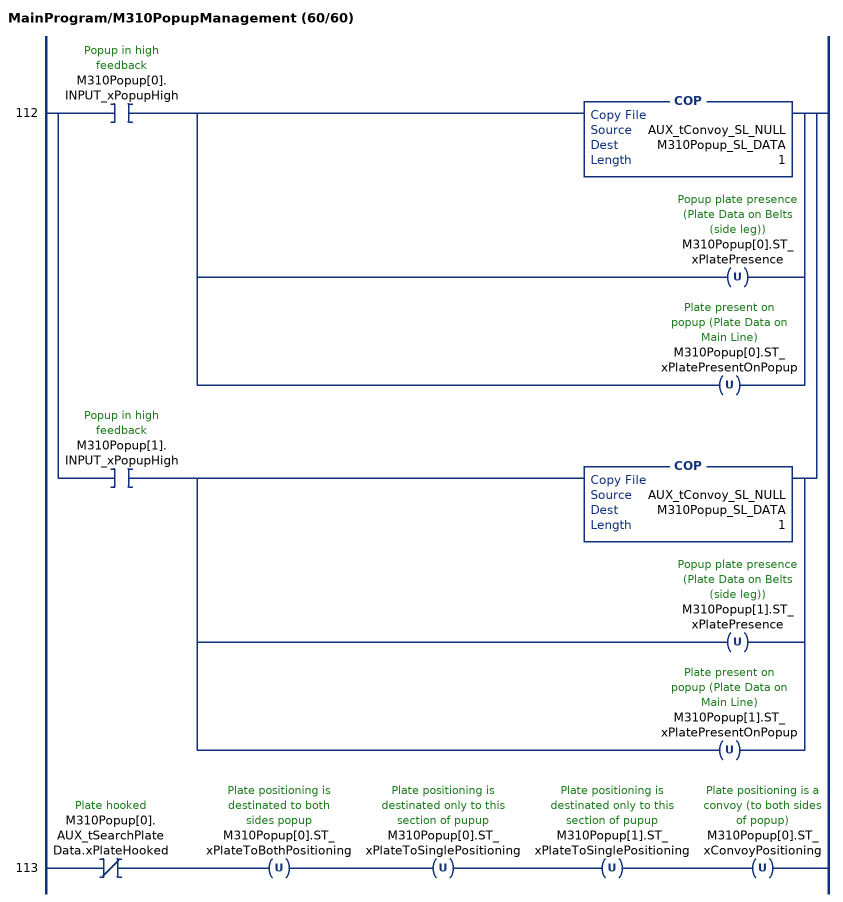
   112: [XIC(M310Popup[0].INPUT_xPopupHigh) [COP(AUX_tConvoy_SL_NULL,M310Popup_SL_DATA,1) ,OTU(M310Popup[0].ST_xPlatePresence) ,OTU(M310Popup[0].ST_xPlatePresentOnPopup) ] ,XIC(M310Popup[1].INPUT_xPopupHigh) [COP(AUX_tConvoy_SL_NULL,M310Popup_SL_DATA,1) ,OTU(M310Popup[1].ST_xPlatePresence) ,OTU(M310Popup[1].ST_xPlatePresentOnPopup) ] ];
   113: XIO(M310Popup[0].AUX_tSearchPlateData.xPlateHooked)OTU(M310Popup[0].ST_xPlateToBothPositioning)OTU(M310Popup[0].ST_xPlateToSinglePositioning)OTU(M310Popup[1].ST_xPlateToSinglePositioning)OTU(M310Popup[0].ST_xConvoyPositioning);
END_ROUTINE

ROUTINE M311_Alarm   (* ladder *)
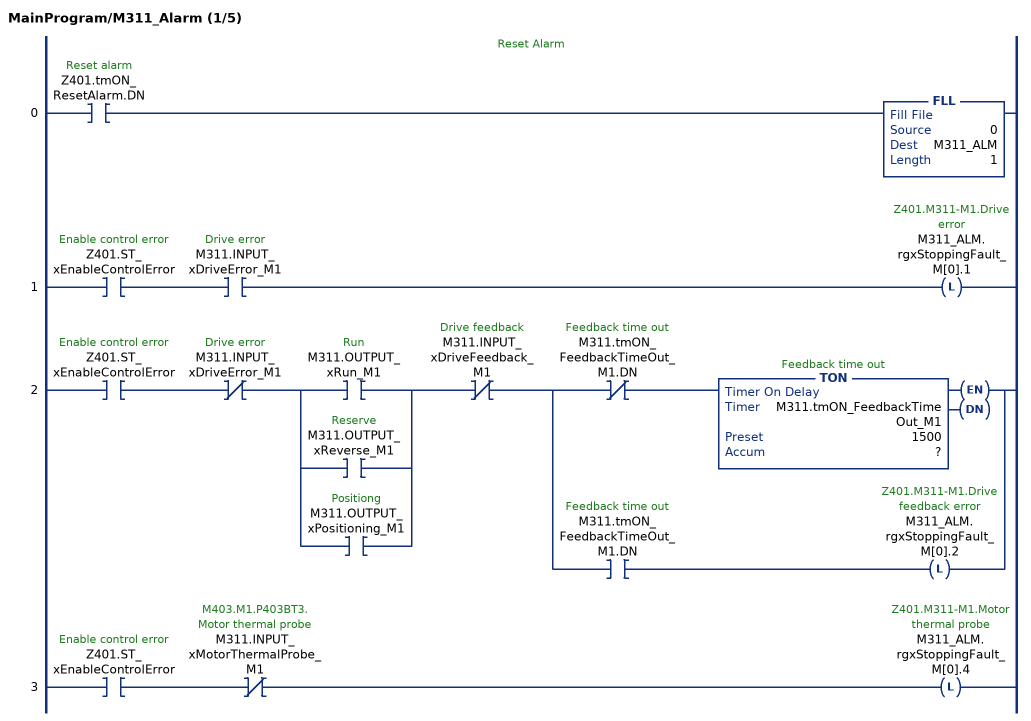
   // Reset Alarm
   0: XIC(Z401.tmON_ResetAlarm.DN)FLL(0,M311_ALM,1);
   1: XIC(Z401.ST_xEnableControlError)XIC(M311.INPUT_xDriveError_M1)OTL(M311_ALM.rgxStoppingFault_M[0].1);
   2: XIC(Z401.ST_xEnableControlError)XIO(M311.INPUT_xDriveError_M1)[XIC(M311.OUTPUT_xRun_M1) ,XIC(M311.OUTPUT_xReverse_M1) ,XIC(M311.OUTPUT_xPositioning_M1) ]XIO(M311.INPUT_xDriveFeedback_M1)[XIO(M311.tmON_FeedbackTimeOut_M1.DN) TON(M311.tmON_FeedbackTimeOut_M1,?,?) ,XIC(M311.tmON_FeedbackTimeOut_M1.DN) OTL(M311_ALM.rgxStoppingFault_M[0].2) ];
   3: XIC(Z401.ST_xEnableControlError)XIO(M311.INPUT_xMotorThermalProbe_M1)OTL(M311_ALM.rgxStoppingFault_M[0].4);
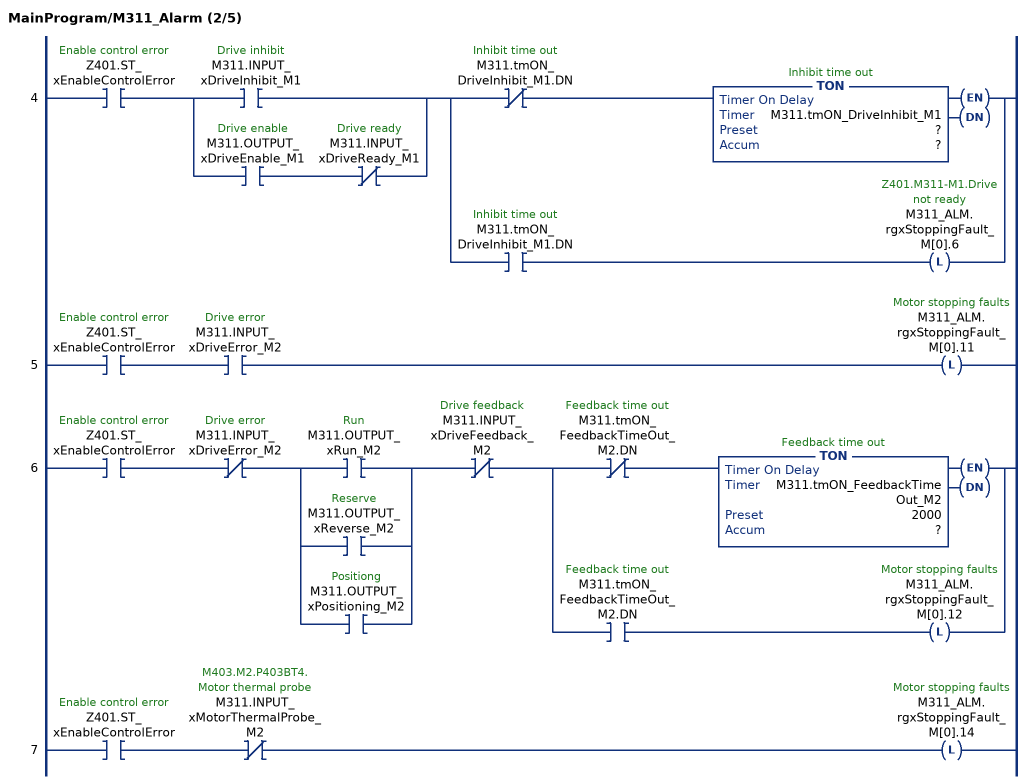
   4: XIC(Z401.ST_xEnableControlError)[XIC(M311.INPUT_xDriveInhibit_M1) ,XIC(M311.OUTPUT_xDriveEnable_M1) XIO(M311.INPUT_xDriveReady_M1) ][XIO(M311.tmON_DriveInhibit_M1.DN) TON(M311.tmON_DriveInhibit_M1,?,?) ,XIC(M311.tmON_DriveInhibit_M1.DN) OTL(M311_ALM.rgxStoppingFault_M[0].6) ];
   5: XIC(Z401.ST_xEnableControlError)XIC(M311.INPUT_xDriveError_M2)OTL(M311_ALM.rgxStoppingFault_M[0].11);
   6: XIC(Z401.ST_xEnableControlError)XIO(M311.INPUT_xDriveError_M2)[XIC(M311.OUTPUT_xRun_M2) ,XIC(M311.OUTPUT_xReverse_M2) ,XIC(M311.OUTPUT_xPositioning_M2) ]XIO(M311.INPUT_xDriveFeedback_M2)[XIO(M311.tmON_FeedbackTimeOut_M2.DN) TON(M311.tmON_FeedbackTimeOut_M2,?,?) ,XIC(M311.tmON_FeedbackTimeOut_M2.DN) OTL(M311_ALM.rgxStoppingFault_M[0].12) ];
   7: XIC(Z401.ST_xEnableControlError)XIO(M311.INPUT_xMotorThermalProbe_M2)OTL(M311_ALM.rgxStoppingFault_M[0].14);
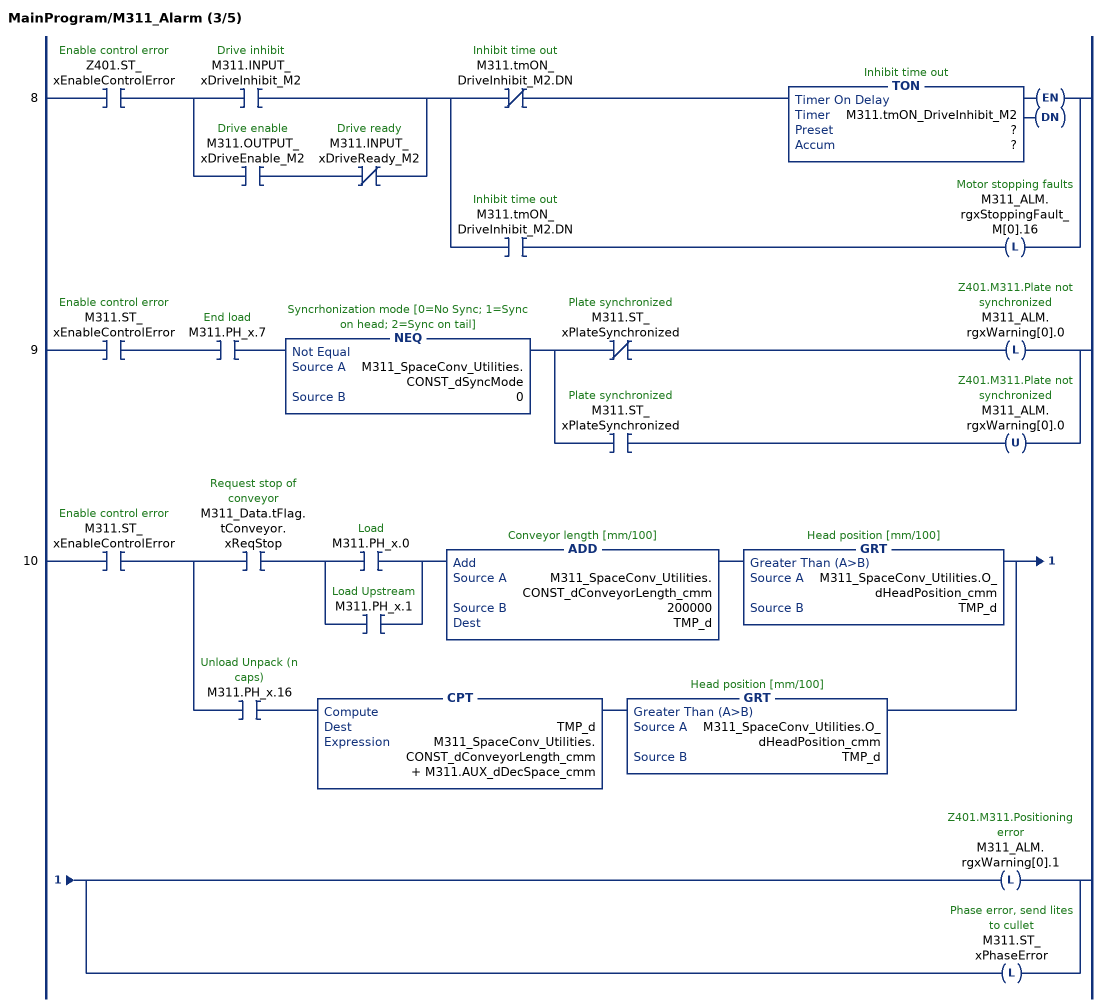
   8: XIC(Z401.ST_xEnableControlError)[XIC(M311.INPUT_xDriveInhibit_M2) ,XIC(M311.OUTPUT_xDriveEnable_M2) XIO(M311.INPUT_xDriveReady_M2) ][XIO(M311.tmON_DriveInhibit_M2.DN) TON(M311.tmON_DriveInhibit_M2,?,?) ,XIC(M311.tmON_DriveInhibit_M2.DN) OTL(M311_ALM.rgxStoppingFault_M[0].16) ];
   9: XIC(M311.ST_xEnableControlError)XIC(M311.PH_x.7)NEQ(M311_SpaceConv_Utilities.CONST_dSyncMode,0)[XIO(M311.ST_xPlateSynchronized) OTL(M311_ALM.rgxWarning[0].0) ,XIC(M311.ST_xPlateSynchronized) OTU(M311_ALM.rgxWarning[0].0) ];
   10: XIC(M311.ST_xEnableControlError)[XIC(M311_Data.tFlag.tConveyor.xReqStop) [XIC(M311.PH_x.0) ,XIC(M311.PH_x.1) ] ADD(M311_SpaceConv_Utilities.CONST_dConveyorLength_cmm,200000,TMP_d) GRT(M311_SpaceConv_Utilities.O_dHeadPosition_cmm,TMP_d) ,XIC(M311.PH_x.16) CPT(TMP_d,M311_SpaceConv_Utilities.CONST_dConveyorLength_cmm + M311.AUX_dDecSpace_cmm) GRT(M311_SpaceConv_Utilities.O_dHeadPosition_cmm,TMP_d) ][OTL(M311_ALM.rgxWarning[0].1) ,OTL(M311.ST_xPhaseError) ];
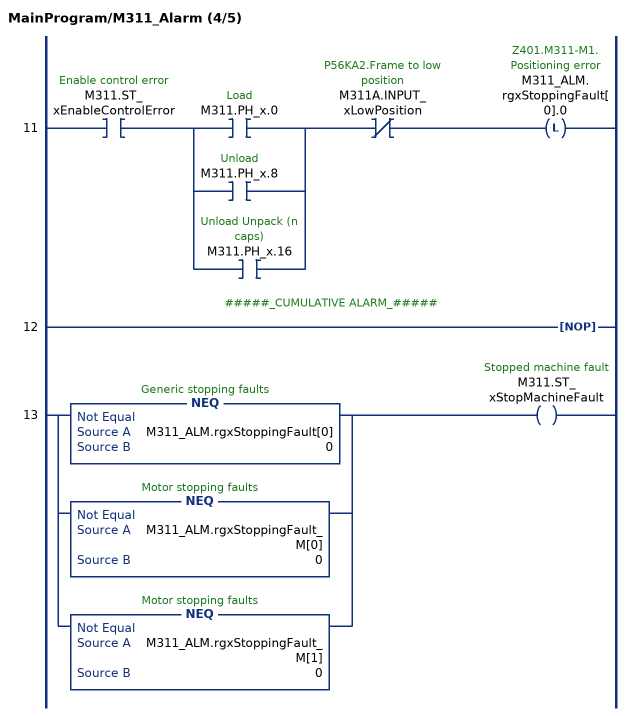
   11: XIC(M311.ST_xEnableControlError)[XIC(M311.PH_x.0) ,XIC(M311.PH_x.8) ,XIC(M311.PH_x.16) ]XIO(M311A.INPUT_xLowPosition)OTL(M311_ALM.rgxStoppingFault[0].0);
   // #####_CUMULATIVE ALARM_#####
   12: NOP();
   13: [NEQ(M311_ALM.rgxStoppingFault[0],0) ,NEQ(M311_ALM.rgxStoppingFault_M[0],0) ,NEQ(M311_ALM.rgxStoppingFault_M[1],0) ]OTE(M311.ST_xStopMachineFault);
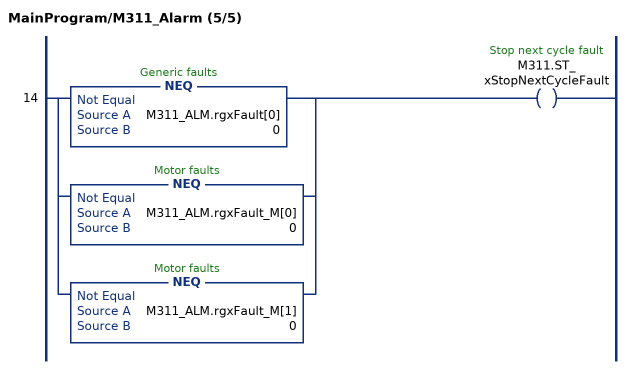
   14: [NEQ(M311_ALM.rgxFault[0],0) ,NEQ(M311_ALM.rgxFault_M[0],0) ,NEQ(M311_ALM.rgxFault_M[1],0) ]OTE(M311.ST_xStopNextCycleFault);
END_ROUTINE

ROUTINE M311_Logic   (* ladder *)
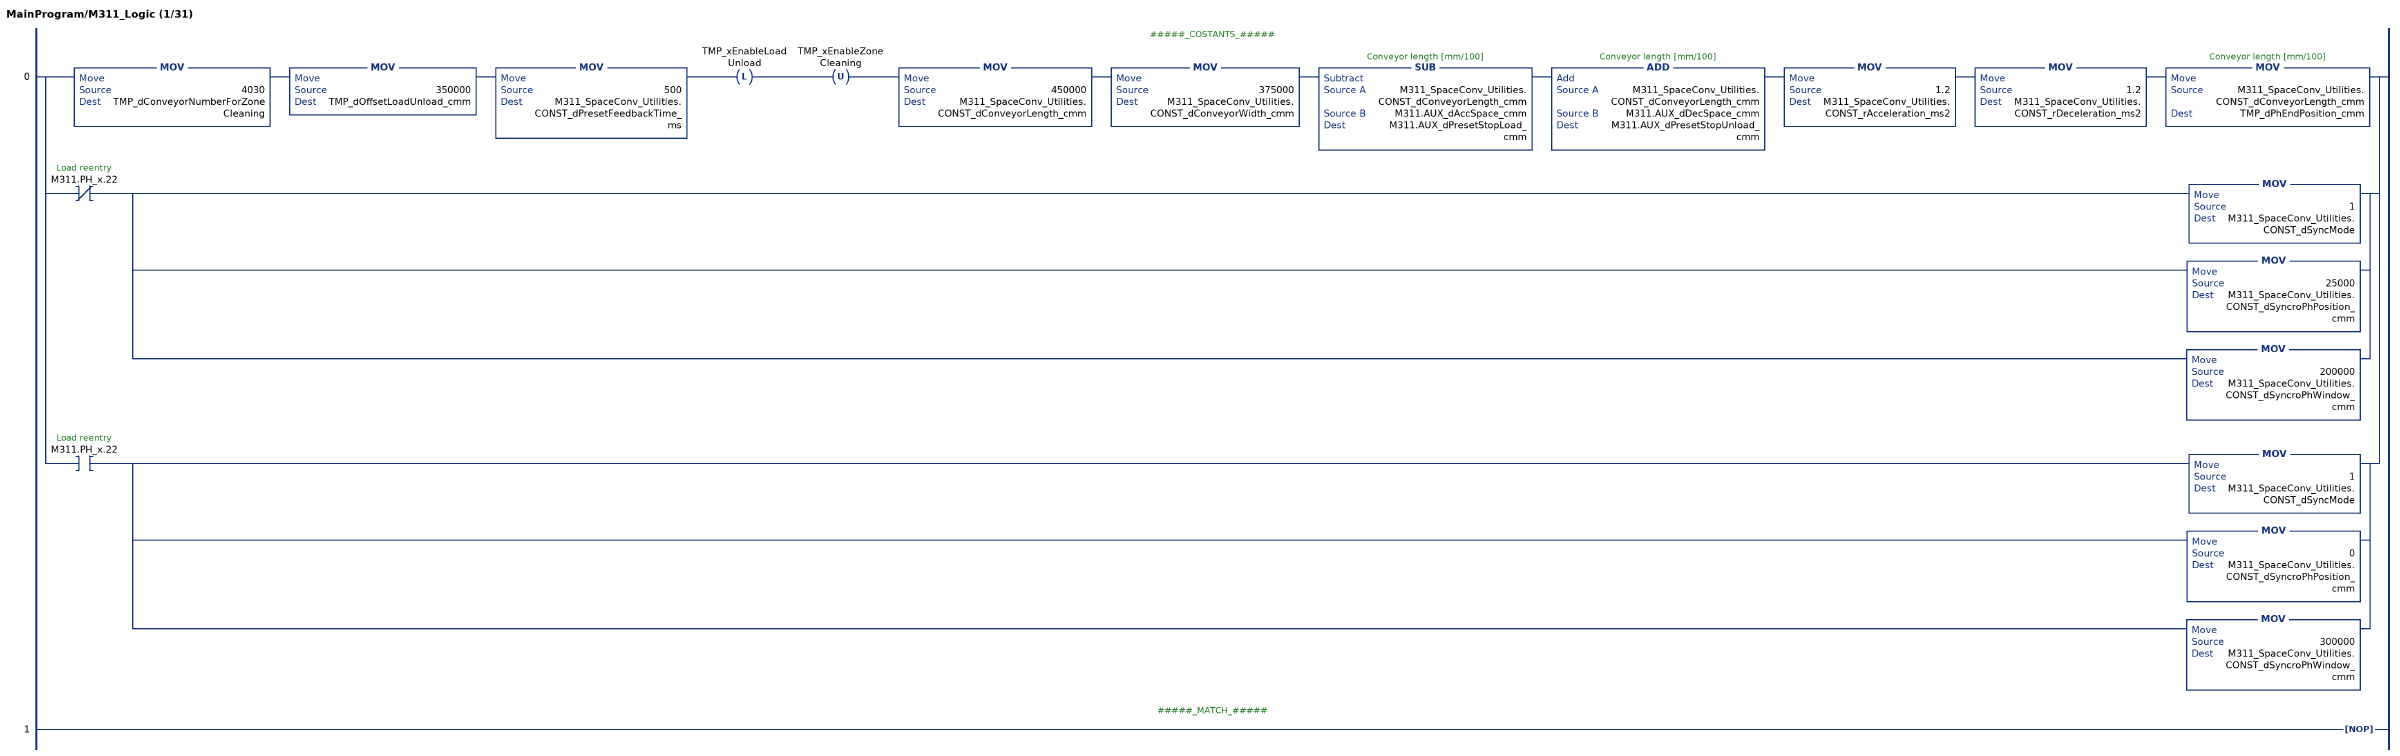
   // #####_COSTANTS_#####
   0: [MOV(4030,TMP_dConveyorNumberForZoneCleaning) MOV(350000,TMP_dOffsetLoadUnload_cmm) MOV(500,M311_SpaceConv_Utilities.CONST_dPresetFeedbackTime_ms) OTL(TMP_xEnableLoadUnload) OTU(TMP_xEnableZoneCleaning) MOV(450000,M311_SpaceConv_Utilities.CONST_dConveyorLength_cmm) MOV(375000,M311_SpaceConv_Utilities.CONST_dConveyorWidth_cmm) SUB(M311_SpaceConv_Utilities.CONST_dConveyorLength_cmm,M311.AUX_dAccSpace_cmm,M311.AUX_dPresetStopLoad_cmm) ADD(M311_SpaceConv_Utilities.CONST_dConveyorLength_cmm,M311.AUX_dDecSpace_cmm,M311.AUX_dPresetStopUnload_cmm) MOV(1.2,M311_SpaceConv_Utilities.CONST_rAcceleration_ms2) MOV(1.2,M311_SpaceConv_Utilities.CONST_rDeceleration_ms2) MOV(M311_SpaceConv_Utilities.CONST_dConveyorLength_cmm,TMP_dPhEndPosition_cmm) ,XIO(M311.PH_x.22) [MOV(1,M311_SpaceConv_Utilities.CONST_dSyncMode) ,MOV(25000,M311_SpaceConv_Utilities.CONST_dSyncroPhPosition_cmm) ,MOV(200000,M311_SpaceConv_Utilities.CONST_dSyncroPhWindow_cmm) ] ,XIC(M311.PH_x.22) [MOV(1,M311_SpaceConv_Utilities.CONST_dSyncMode) ,MOV(0,M311_SpaceConv_Utilities.CONST_dSyncroPhPosition_cmm) ,MOV(300000,M311_SpaceConv_Utilities.CONST_dSyncroPhWindow_cmm) ] ];
   // #####_MATCH_#####
   1: NOP();
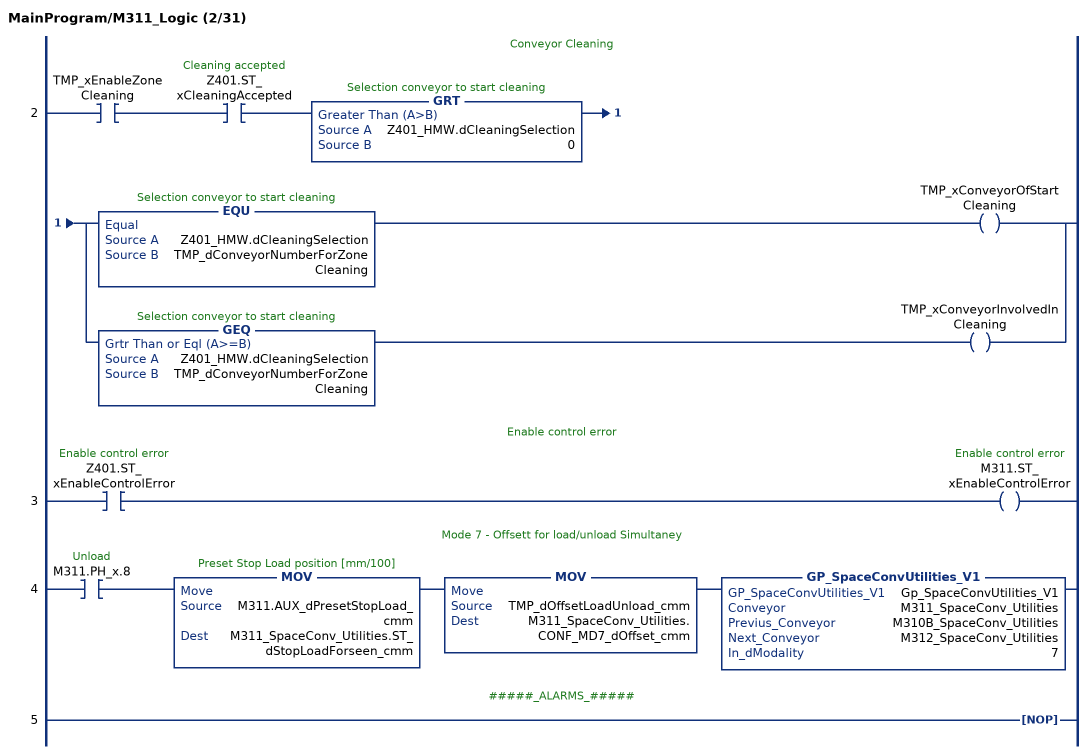
   // Conveyor Cleaning
   2: XIC(TMP_xEnableZoneCleaning)XIC(Z401.ST_xCleaningAccepted)GRT(Z401_HMW.dCleaningSelection,0)[EQU(Z401_HMW.dCleaningSelection,TMP_dConveyorNumberForZoneCleaning) OTE(TMP_xConveyorOfStartCleaning) ,GEQ(Z401_HMW.dCleaningSelection,TMP_dConveyorNumberForZoneCleaning) OTE(TMP_xConveyorInvolvedInCleaning) ];
   // Enable control error
   3: XIC(Z401.ST_xEnableControlError)OTE(M311.ST_xEnableControlError);
   // Mode 7 - Offsett for load/unload Simultaney
   4: XIC(M311.PH_x.8)MOV(M311.AUX_dPresetStopLoad_cmm,M311_SpaceConv_Utilities.ST_dStopLoadForseen_cmm)MOV(TMP_dOffsetLoadUnload_cmm,M311_SpaceConv_Utilities.CONF_MD7_dOffset_cmm)GP_SpaceConvUtilities_V1(Gp_SpaceConvUtilities_V1,M311_SpaceConv_Utilities,M310B_SpaceConv_Utilities,M312_SpaceConv_Utilities,7);
   // #####_ALARMS_#####
   5: NOP();
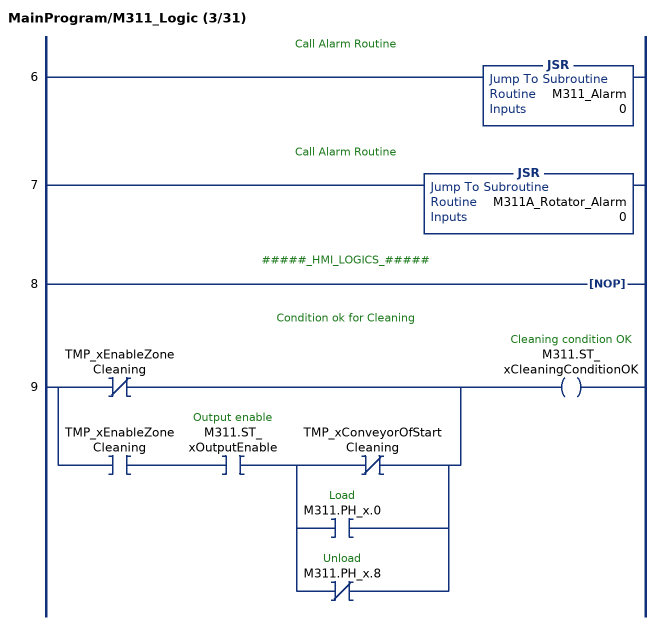
   // Call Alarm Routine
   6: JSR(M311_Alarm,0);
   // Call Alarm Routine
   7: JSR(M311A_Rotator_Alarm,0);
   // #####_HMI_LOGICS_#####
   8: NOP();
   // Condition ok for Cleaning
   9: [XIO(TMP_xEnableZoneCleaning) ,XIC(TMP_xEnableZoneCleaning) XIC(M311.ST_xOutputEnable) [XIO(TMP_xConveyorOfStartCleaning) ,XIC(M311.PH_x.0) ,XIO(M311.PH_x.8) ] ]OTE(M311.ST_xCleaningConditionOK);
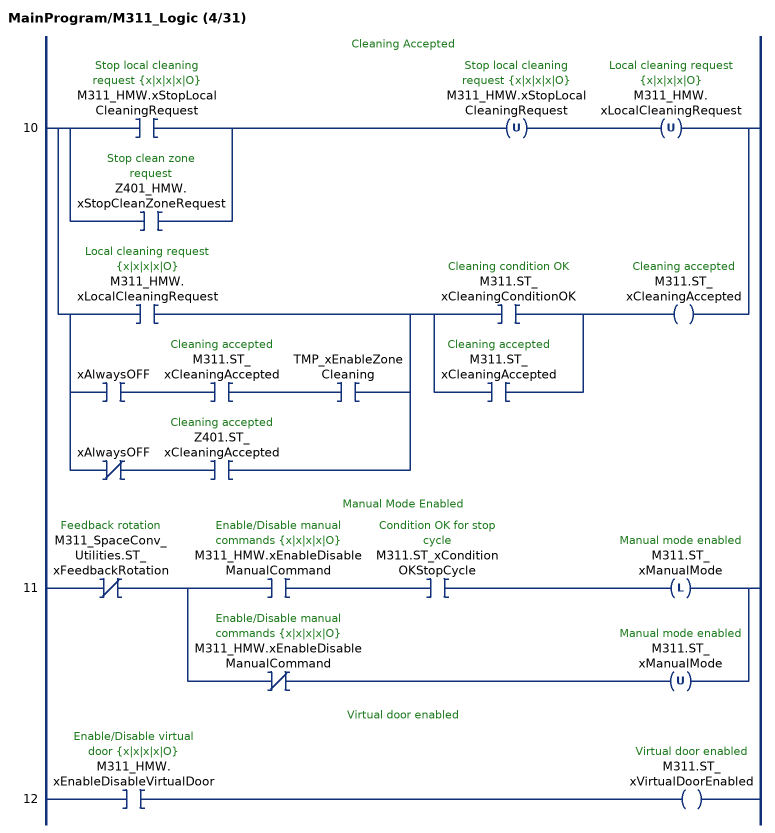
   // Cleaning Accepted
   10: [[XIC(M311_HMW.xStopLocalCleaningRequest) ,XIC(Z401_HMW.xStopCleanZoneRequest) ] OTU(M311_HMW.xStopLocalCleaningRequest) OTU(M311_HMW.xLocalCleaningRequest) ,[XIC(M311_HMW.xLocalCleaningRequest) ,XIC(xAlwaysOFF) XIC(M311.ST_xCleaningAccepted) XIC(TMP_xEnableZoneCleaning) ,XIO(xAlwaysOFF) XIC(Z401.ST_xCleaningAccepted) ] [XIC(M311.ST_xCleaningConditionOK) ,XIC(M311.ST_xCleaningAccepted) ] OTE(M311.ST_xCleaningAccepted) ];
   // Manual Mode Enabled
   11: XIO(M311_SpaceConv_Utilities.ST_xFeedbackRotation)[XIC(M311_HMW.xEnableDisableManualCommand) XIC(M311.ST_xConditionOKStopCycle) OTL(M311.ST_xManualMode) ,XIO(M311_HMW.xEnableDisableManualCommand) OTU(M311.ST_xManualMode) ];
   // Virtual door enabled
   12: XIC(M311_HMW.xEnableDisableVirtualDoor)OTE(M311.ST_xVirtualDoorEnabled);
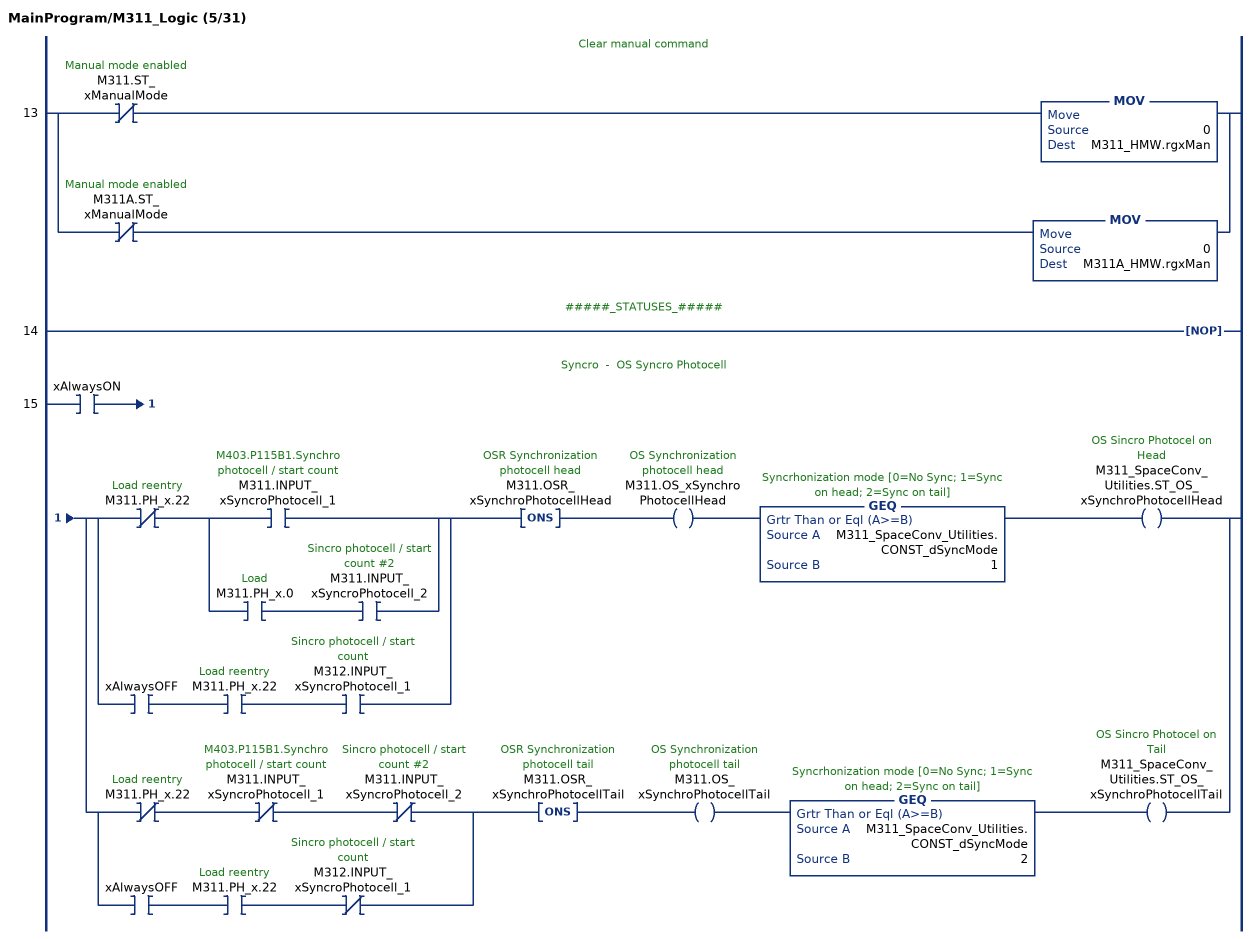
   // Clear manual command
   13: [XIO(M311.ST_xManualMode) MOV(0,M311_HMW.rgxMan) ,XIO(M311A.ST_xManualMode) MOV(0,M311A_HMW.rgxMan) ];
   // #####_STATUSES_#####
   14: NOP();
   // Syncro  -  OS Syncro Photocell
   15: XIC(xAlwaysON)[[XIO(M311.PH_x.22) [XIC(M311.INPUT_xSyncroPhotocell_1) ,XIC(M311.PH_x.0) XIC(M311.INPUT_xSyncroPhotocell_2) ] ,XIC(xAlwaysOFF) XIC(M311.PH_x.22) XIC(M312.INPUT_xSyncroPhotocell_1) ] ONS(M311.OSR_xSynchroPhotocellHead) OTE(M311.OS_xSynchroPhotocellHead) GEQ(M311_SpaceConv_Utilities.CONST_dSyncMode,1) OTE(M311_SpaceConv_Utilities.ST_OS_xSynchroPhotocellHead) ,[XIO(M311.PH_x.22) XIO(M311.INPUT_xSyncroPhotocell_1) XIO(M311.INPUT_xSyncroPhotocell_2) ,XIC(xAlwaysOFF) XIC(M311.PH_x.22) XIO(M312.INPUT_xSyncroPhotocell_1) ] ONS(M311.OSR_xSynchroPhotocellTail) OTE(M311.OS_xSynchroPhotocellTail) GEQ(M311_SpaceConv_Utilities.CONST_dSyncMode,2) OTE(M311_SpaceConv_Utilities.ST_OS_xSynchroPhotocellTail) ];
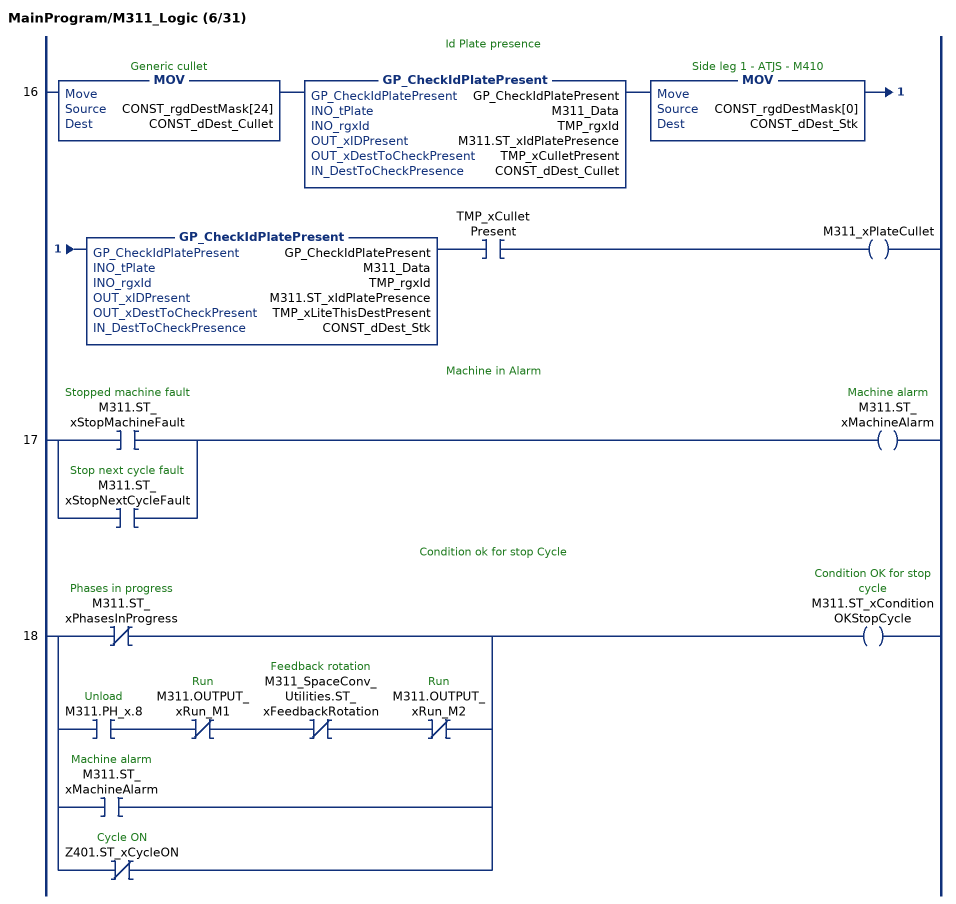
   // Id Plate presence
   16: MOV(CONST_rgdDestMask[24],CONST_dDest_Cullet)GP_CheckIdPlatePresent(GP_CheckIdPlatePresent,M311_Data,TMP_rgxId,M311.ST_xIdPlatePresence,TMP_xCulletPresent,CONST_dDest_Cullet)MOV(CONST_rgdDestMask[0],CONST_dDest_Stk)GP_CheckIdPlatePresent(GP_CheckIdPlatePresent,M311_Data,TMP_rgxId,M311.ST_xIdPlatePresence,TMP_xLiteThisDestPresent,CONST_dDest_Stk)XIC(TMP_xCulletPresent)OTE(M311_xPlateCullet);
   // Machine in Alarm
   17: [XIC(M311.ST_xStopMachineFault) ,XIC(M311.ST_xStopNextCycleFault) ]OTE(M311.ST_xMachineAlarm);
   // Condition ok for stop Cycle
   18: [XIO(M311.ST_xPhasesInProgress) ,XIC(M311.PH_x.8) XIO(M311.OUTPUT_xRun_M1) XIO(M311_SpaceConv_Utilities.ST_xFeedbackRotation) XIO(M311.OUTPUT_xRun_M2) ,XIC(M311.ST_xMachineAlarm) ,XIO(Z401.ST_xCycleON) ]OTE(M311.ST_xConditionOKStopCycle);
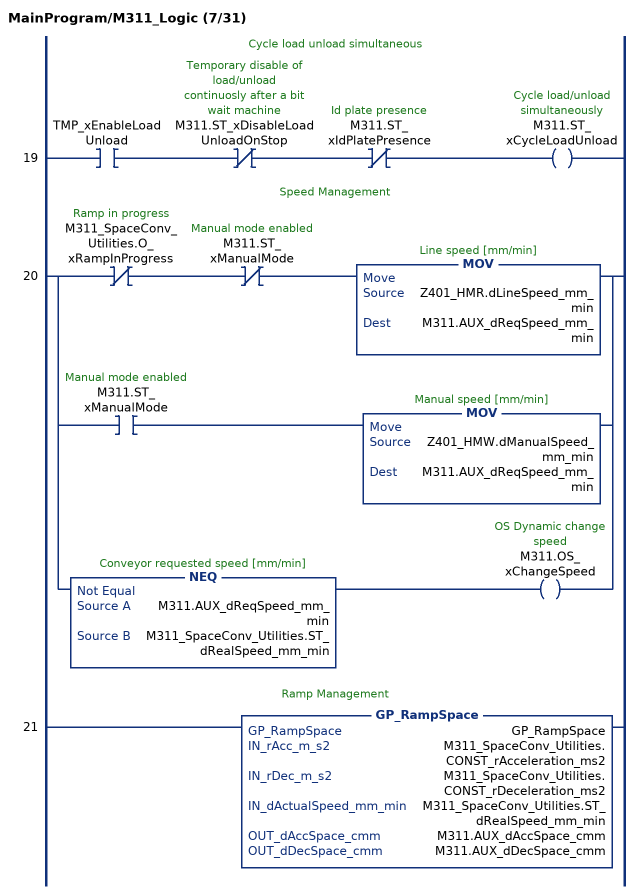
   // Cycle load unload simultaneous
   19: XIC(TMP_xEnableLoadUnload)XIO(M311.ST_xDisableLoadUnloadOnStop)XIO(M311.ST_xIdPlatePresence)OTE(M311.ST_xCycleLoadUnload);
   // Speed Management
   20: [XIO(M311_SpaceConv_Utilities.O_xRampInProgress) XIO(M311.ST_xManualMode) MOV(Z401_HMR.dLineSpeed_mm_min,M311.AUX_dReqSpeed_mm_min) ,XIC(M311.ST_xManualMode) MOV(Z401_HMW.dManualSpeed_mm_min,M311.AUX_dReqSpeed_mm_min) ,NEQ(M311.AUX_dReqSpeed_mm_min,M311_SpaceConv_Utilities.ST_dRealSpeed_mm_min) OTE(M311.OS_xChangeSpeed) ];
   // Ramp Management
   21: GP_RampSpace(GP_RampSpace,M311_SpaceConv_Utilities.CONST_rAcceleration_ms2,M311_SpaceConv_Utilities.CONST_rDeceleration_ms2,M311_SpaceConv_Utilities.ST_dRealSpeed_mm_min,M311.AUX_dAccSpace_cmm,M311.AUX_dDecSpace_cmm);
